D3525:=ComConveyorIO701102.o_iRequestPLCPC; 
D3526:=ComConveyorIO701102.o_iForceInportPLCPC;
D3527:=ComConveyorIO701102.o_iFolderNumberPLCPC;
D3528:=ComConveyorIO701102.o_iEmptyPLCPC;
D3530:=ComConveyorIO701102.o_iReadWriteFlagPLCPC; 
D3531:=ComConveyorIO701102.o_iDeviceStatusPLCPC; 
D3532:=ComConveyorIO701102.o_iTaskIDPLCPC; 
D3533:=ComConveyorIO701102.o_iProductIDPLCPC;
ComConveyorIO701102.i_xExportConveyor:=1;
ComConveyorIO701102.i_xExtraCondition:=ConveyorIO70159.xEmpty AND NOT ConveyorIO70159.xCWPresent AND NOT ConveyorIO701102.xCWPresent;*)
(*F5出库站台1*)
ComConveyorIO70159.i_iResponsPCPLC:=D2540; 
ComConveyorIO70159.i_iTypeInfoPCPLC:=D2541;
ComConveyorIO70159.i_iReadWriteFlagPCPLC:=D2545; 
ComConveyorIO70159.i_iTaskProcessFlagPCPLC:=D2546; 
ComConveyorIO70159.i_iCommandPCPLC:=D2547; 
ComConveyorIO70159.i_iTaskIDPCPLC:=D2548; 
DMOV(TRUE,D2549,ComConveyorIO70159.i_diDestinationDevicePCPLC); 
ComConveyorIO70159.i_iProductIDPCPLC:=D2551;
D3540:=ComConveyorIO70159.o_iRequestPLCPC; 
D3541:=ComConveyorIO70159.o_iForceInportPLCPC;
D3542:=ComConveyorIO70159.o_iFolderNumberPLCPC;
D3543:=ComConveyorIO70159.o_iEmptyPLCPC;
D3545:=ComConveyorIO70159.o_iReadWriteFlagPLCPC; 
D3546:=ComConveyorIO70159.o_iDeviceStatusPLCPC; 
D3547:=ComConveyorIO70159.o_iTaskIDPLCPC; 
D3548:=ComConveyorIO70159.o_iProductIDPLCPC;
ComConveyorIO70159.i_xExportConveyor:=1;
ComConveyorIO70159.i_xExtraCondition:=ConveyorIO701102.xEmpty AND NOT ConveyorIO70159.xCWPresent AND NOT ConveyorIO701102.xCWPresent;
(*F6出库站台1*)
ComConveyorIO701120.i_iResponsPCPLC:=D2555; 
ComConveyorIO701120.i_iTypeInfoPCPLC:=D2556;
ComConveyorIO701120.i_iReadWriteFlagPCPLC:=D2560; 
ComConveyorIO701120.i_iTaskProcessFlagPCPLC:=D2561; 
ComConveyorIO701120.i_iCommandPCPLC:=D2562; 
ComConveyorIO701120.i_iTaskIDPCPLC:=D2563; 
DMOV(TRUE,D2564,ComConveyorIO701120.i_diDestinationDevicePCPLC); 
ComConveyorIO701120.i_iProductIDPCPLC:=D2566;
D3555:=ComConveyorIO701120.o_iRequestPLCPC; 
D3556:=ComConveyorIO701120.o_iForceInportPLCPC;
D3557:=ComConveyorIO701120.o_iFolderNumberPLCPC;
D3558:=ComConveyorIO701120.o_iEmptyPLCPC;
D3560:=ComConveyorIO701120.o_iReadWriteFlagPLCPC; 
D3561:=ComConveyorIO701120.o_iDeviceStatusPLCPC; 
D3562:=ComConveyorIO701120.o_iTaskIDPLCPC; 
D3563:=ComConveyorIO701120.o_iProductIDPLCPC;
ComConveyorIO701120.i_xExportConveyor:=1;
ComConveyorIO701120.i_xExtraCondition:=ConveyorIO701119.xEmpty AND NOT ConveyorIO701119.xCWPresent AND NOT ConveyorIO701120.xCWPresent;
(*
ComConveyorIO701119.i_iResponsPCPLC:=D2570; 
ComConveyorIO701119.i_iTypeInfoPCPLC:=D2571;
ComConveyorIO701119.i_iReadWriteFlagPCPLC:=D2575; 
ComConveyorIO701119.i_iTaskProcessFlagPCPLC:=D2576; 
ComConveyorIO701119.i_iCommandPCPLC:=D2577; 
ComConveyorIO701119.i_iTaskIDPCPLC:=D2578; 
DMOV(TRUE,D2579,ComConveyorIO701119.i_diDestinationDevicePCPLC); 
ComConveyorIO701119.i_iProductIDPCPLC:=D2581;
D3570:=ComConveyorIO701119.o_iRequestPLCPC; 
D3571:=ComConveyorIO701119.o_iForceInportPLCPC;
D3572:=ComConveyorIO701119.o_iFolderNumberPLCPC;
D3573:=ComConveyorIO701119.o_iEmptyPLCPC;
D3575:=ComConveyorIO701119.o_iReadWriteFlagPLCPC; 
D3576:=ComConveyorIO701119.o_iDeviceStatusPLCPC; 
D3577:=ComConveyorIO701119.o_iTaskIDPLCPC; 
D3578:=ComConveyorIO701119.o_iProductIDPLCPC;
ComConveyorIO701119.i_xExportConveyor:=1;*)
(*F1空框入库站台2*)
ComConveyorIO701105.i_iTypeInfoPCPLC:=D2616;
ComConveyorIO701105.i_iReadWriteFlagPCPLC:=D2620; 
ComConveyorIO701105.i_iTaskProcessFlagPCPLC:=D2621; 
ComConveyorIO701105.i_iCommandPCPLC:=D2622; 
ComConveyorIO701105.i_iTaskIDPCPLC:=D2623; 
DMOV(TRUE,D2624,ComConveyorIO701105.i_diDestinationDevicePCPLC); 
ComConveyorIO701105.i_iProductIDPCPLC:=D2626;
D3615:=ComConveyorIO701105.o_iRequestPLCPC; 
D3616:=ComConveyorIO701105.o_iForceInportPLCPC;
D3617:=ComConveyorIO701105.o_iFolderNumberPLCPC;
D3618:=ComConveyorIO701105.o_iEmptyPLCPC;
D3620:=ComConveyorIO701105.o_iReadWriteFlagPLCPC; 
D3621:=ComConveyorIO701105.o_iDeviceStatusPLCPC; 
D3622:=ComConveyorIO701105.o_iTaskIDPLCPC; 
D3623:=ComConveyorIO701105.o_iProductIDPLCPC;
(*F2空框入库站台1*)
ComConveyorIO70113.i_iResponsPCPLC:=D2630; 
ComConveyorIO70113.i_iTypeInfoPCPLC:=D2631;
ComConveyorIO70113.i_iReadWriteFlagPCPLC:=D2635; 
ComConveyorIO70113.i_iTaskProcessFlagPCPLC:=D2636; 
ComConveyorIO70113.i_iCommandPCPLC:=D2637; 
ComConveyorIO70113.i_iTaskIDPCPLC:=D2638; 
DMOV(TRUE,D2639,ComConveyorIO70113.i_diDestinationDevicePCPLC); 
ComConveyorIO70113.i_iProductIDPCPLC:=D2641;
D3630:=ComConveyorIO70113.o_iRequestPLCPC; 
D3631:=ComConveyorIO70113.o_iForceInportPLCPC;
D3632:=ComConveyorIO70113.o_iFolderNumberPLCPC;
D3633:=ComConveyorIO70113.o_iEmptyPLCPC;
D3635:=ComConveyorIO70113.o_iReadWriteFlagPLCPC; 
D3636:=ComConveyorIO70113.o_iDeviceStatusPLCPC; 
D3637:=ComConveyorIO70113.o_iTaskIDPLCPC; 
D3638:=ComConveyorIO70113.o_iProductIDPLCPC;
(*F2空框入库站台2*)
ComConveyorIO701106.i_iResponsPCPLC:=D2645; 
ComConveyorIO701106.i_iTypeInfoPCPLC:=D2646;
ComConveyorIO701106.i_iReadWriteFlagPCPLC:=D2650; 
ComConveyorIO701106.i_iTaskProcessFlagPCPLC:=D2651; 
ComConveyorIO701106.i_iCommandPCPLC:=D2652; 
ComConveyorIO701106.i_iTaskIDPCPLC:=D2653; 
DMOV(TRUE,D2654,ComConveyorIO701106.i_diDestinationDevicePCPLC); 
ComConveyorIO701106.i_iProductIDPCPLC:=D2656;
D3645:=ComConveyorIO701106.o_iRequestPLCPC; 
D3646:=ComConveyorIO701106.o_iForceInportPLCPC;
D3647:=ComConveyorIO701106.o_iFolderNumberPLCPC;
D3648:=ComConveyorIO701106.o_iEmptyPLCPC;
D3650:=ComConveyorIO701106.o_iReadWriteFlagPLCPC; 
D3651:=ComConveyorIO701106.o_iDeviceStatusPLCPC; 
D3652:=ComConveyorIO701106.o_iTaskIDPLCPC; 
D3653:=ComConveyorIO701106.o_iProductIDPLCPC;
(*F1,2入库前主路分流站台*)
ComConveyorIO70114.i_iResponsPCPLC:=D2660; 
ComConveyorIO70114.i_iTypeInfoPCPLC:=D2661;
ComConveyorIO70114.i_iReadWriteFlagPCPLC:=D2665; 
ComConveyorIO70114.i_iTaskProcessFlagPCPLC:=D2666; 
ComConveyorIO70114.i_iCommandPCPLC:=D2667; 
ComConveyorIO70114.i_iTaskIDPCPLC:=D2668; 
DMOV(TRUE,D2669,ComConveyorIO70114.i_diDestinationDevicePCPLC); 
ComConveyorIO70114.i_iProductIDPCPLC:=D2671;
D3660:=ComConveyorIO70114.o_iRequestPLCPC; 
D3661:=ComConveyorIO70114.o_iForceInportPLCPC;
D3662:=ComConveyorIO70114.o_iFolderNumberPLCPC;
D3663:=ComConveyorIO70114.o_iEmptyPLCPC;
D3665:=ComConveyorIO70114.o_iReadWriteFlagPLCPC; 
D3666:=ComConveyorIO70114.o_iDeviceStatusPLCPC; 
D3667:=ComConveyorIO70114.o_iTaskIDPLCPC; 
D3668:=ComConveyorIO70114.o_iProductIDPLCPC;
ComConveyorIO70116.i_iTypeInfoPCPLC:=D2691;
ComConveyorIO70116.i_iReadWriteFlagPCPLC:=D2695; 
ComConveyorIO70116.i_iTaskProcessFlagPCPLC:=D2696; 
ComConveyorIO70116.i_iCommandPCPLC:=D2697; 
ComConveyorIO70116.i_iTaskIDPCPLC:=D2698; 
DMOV(TRUE,D2699,ComConveyorIO70116.i_diDestinationDevicePCPLC); 
ComConveyorIO70116.i_iProductIDPCPLC:=D2701;
D3690:=ComConveyorIO70116.o_iRequestPLCPC; 
D3691:=ComConveyorIO70116.o_iForceInportPLCPC;
D3692:=ComConveyorIO70116.o_iFolderNumberPLCPC;
D3693:=ComConveyorIO70116.o_iEmptyPLCPC;
D3695:=ComConveyorIO70116.o_iReadWriteFlagPLCPC; 
D3696:=ComConveyorIO70116.o_iDeviceStatusPLCPC; 
D3697:=ComConveyorIO70116.o_iTaskIDPLCPC; 
D3698:=ComConveyorIO70116.o_iProductIDPLCPC;
ComConveyorIO70119.i_iResponsPCPLC:=D2705; 
ComConveyorIO70119.i_iTypeInfoPCPLC:=D2706;
ComConveyorIO70119.i_iReadWriteFlagPCPLC:=D2710; 
ComConveyorIO70119.i_iTaskProcessFlagPCPLC:=D2711; 
ComConveyorIO70119.i_iCommandPCPLC:=D2712; 
ComConveyorIO70119.i_iTaskIDPCPLC:=D2713; 
DMOV(TRUE,D2714,ComConveyorIO70119.i_diDestinationDevicePCPLC); 
ComConveyorIO70119.i_iProductIDPCPLC:=D2716;
D3705:=ComConveyorIO70119.o_iRequestPLCPC; 
D3706:=ComConveyorIO70119.o_iForceInportPLCPC;
D3707:=ComConveyorIO70119.o_iFolderNumberPLCPC;
D3708:=ComConveyorIO70119.o_iEmptyPLCPC;
D3710:=ComConveyorIO70119.o_iReadWriteFlagPLCPC; 
D3711:=ComConveyorIO70119.o_iDeviceStatusPLCPC; 
D3712:=ComConveyorIO70119.o_iTaskIDPLCPC; 
D3713:=ComConveyorIO70119.o_iProductIDPLCPC;
ComConveyorIO70120.i_iResponsPCPLC:=D2720; 
ComConveyorIO70120.i_iTypeInfoPCPLC:=D2721;
ComConveyorIO70120.i_iReadWriteFlagPCPLC:=D2725; 
ComConveyorIO70120.i_iTaskProcessFlagPCPLC:=D2726; 
ComConveyorIO70120.i_iCommandPCPLC:=D2727; 
ComConveyorIO70120.i_iTaskIDPCPLC:=D2728; 
DMOV(TRUE,D2729,ComConveyorIO70120.i_diDestinationDevicePCPLC); 
ComConveyorIO70120.i_iProductIDPCPLC:=D2731;
D3720:=ComConveyorIO70120.o_iRequestPLCPC; 
D3721:=ComConveyorIO70120.o_iForceInportPLCPC;
D3722:=ComConveyorIO70120.o_iFolderNumberPLCPC;
D3723:=ComConveyorIO70120.o_iEmptyPLCPC;
D3725:=ComConveyorIO70120.o_iReadWriteFlagPLCPC; 
D3726:=ComConveyorIO70120.o_iDeviceStatusPLCPC; 
D3727:=ComConveyorIO70120.o_iTaskIDPLCPC; 
D3728:=ComConveyorIO70120.o_iProductIDPLCPC;
ComConveyorIO701107.i_iResponsPCPLC:=D2735; 
ComConveyorIO701107.i_iTypeInfoPCPLC:=D2736;
ComConveyorIO701107.i_iReadWriteFlagPCPLC:=D2740; 
ComConveyorIO701107.i_iTaskProcessFlagPCPLC:=D2741; 
ComConveyorIO701107.i_iCommandPCPLC:=D2742; 
ComConveyorIO701107.i_iTaskIDPCPLC:=D2743; 
DMOV(TRUE,D2744,ComConveyorIO701107.i_diDestinationDevicePCPLC); 
ComConveyorIO701107.i_iProductIDPCPLC:=D2746;
D3735:=ComConveyorIO701107.o_iRequestPLCPC; 
D3736:=ComConveyorIO701107.o_iForceInportPLCPC;
D3737:=ComConveyorIO701107.o_iFolderNumberPLCPC;
D3738:=ComConveyorIO701107.o_iEmptyPLCPC;
D3740:=ComConveyorIO701107.o_iReadWriteFlagPLCPC; 
D3741:=ComConveyorIO701107.o_iDeviceStatusPLCPC; 
D3742:=ComConveyorIO701107.o_iTaskIDPLCPC; 
D3743:=ComConveyorIO701107.o_iProductIDPLCPC;
ComConveyorIO70121.i_iResponsPCPLC:=D2750; 
ComConveyorIO70121.i_iTypeInfoPCPLC:=D2751;
ComConveyorIO70121.i_iReadWriteFlagPCPLC:=D2755; 
ComConveyorIO70121.i_iTaskProcessFlagPCPLC:=D2756; 
ComConveyorIO70121.i_iCommandPCPLC:=D2757; 
ComConveyorIO70121.i_iTaskIDPCPLC:=D2758; 
DMOV(TRUE,D2759,ComConveyorIO70121.i_diDestinationDevicePCPLC); 
ComConveyorIO70121.i_iProductIDPCPLC:=D2761;
D3750:=ComConveyorIO70121.o_iRequestPLCPC; 
D3751:=ComConveyorIO70121.o_iForceInportPLCPC;
D3752:=ComConveyorIO70121.o_iFolderNumberPLCPC;
D3753:=ComConveyorIO70121.o_iEmptyPLCPC;
D3755:=ComConveyorIO70121.o_iReadWriteFlagPLCPC; 
D3756:=ComConveyorIO70121.o_iDeviceStatusPLCPC; 
D3757:=ComConveyorIO70121.o_iTaskIDPLCPC; 
D3758:=ComConveyorIO70121.o_iProductIDPLCPC;
ComConveyorIO701108.i_iResponsPCPLC:=D2765; 
ComConveyorIO701108.i_iTypeInfoPCPLC:=D2766;
ComConveyorIO701108.i_iReadWriteFlagPCPLC:=D2770; 
ComConveyorIO701108.i_iTaskProcessFlagPCPLC:=D2771; 
ComConveyorIO701108.i_iCommandPCPLC:=D2772; 
ComConveyorIO701108.i_iTaskIDPCPLC:=D2773; 
DMOV(TRUE,D2774,ComConveyorIO701108.i_diDestinationDevicePCPLC); 
ComConveyorIO701108.i_iProductIDPCPLC:=D2776;
D3765:=ComConveyorIO701108.o_iRequestPLCPC; 
D3766:=ComConveyorIO701108.o_iForceInportPLCPC;
D3767:=ComConveyorIO701108.o_iFolderNumberPLCPC;
D3768:=ComConveyorIO701108.o_iEmptyPLCPC;
D3770:=ComConveyorIO701108.o_iReadWriteFlagPLCPC; 
D3771:=ComConveyorIO701108.o_iDeviceStatusPLCPC; 
D3772:=ComConveyorIO701108.o_iTaskIDPLCPC; 
D3773:=ComConveyorIO701108.o_iProductIDPLCPC;
ComConveyorIO70122.i_iResponsPCPLC:=D2780; 
ComConveyorIO70122.i_iTypeInfoPCPLC:=D2781;
ComConveyorIO70122.i_iReadWriteFlagPCPLC:=D2785; 
ComConveyorIO70122.i_iTaskProcessFlagPCPLC:=D2786; 
ComConveyorIO70122.i_iCommandPCPLC:=D2787; 
ComConveyorIO70122.i_iTaskIDPCPLC:=D2788; 
DMOV(TRUE,D2789,ComConveyorIO70122.i_diDestinationDevicePCPLC); 
ComConveyorIO70122.i_iProductIDPCPLC:=D2791;
D3780:=ComConveyorIO70122.o_iRequestPLCPC; 
D3781:=ComConveyorIO70122.o_iForceInportPLCPC;
D3782:=ComConveyorIO70122.o_iFolderNumberPLCPC;
D3783:=ComConveyorIO70122.o_iEmptyPLCPC;
D3785:=ComConveyorIO70122.o_iReadWriteFlagPLCPC; 
D3786:=ComConveyorIO70122.o_iDeviceStatusPLCPC; 
D3787:=ComConveyorIO70122.o_iTaskIDPLCPC; 
D3788:=ComConveyorIO70122.o_iProductIDPLCPC;
ComConveyorIO70124.i_iResponsPCPLC:=D2795; 
ComConveyorIO70124.i_iTypeInfoPCPLC:=D2796;
ComConveyorIO70124.i_iReadWriteFlagPCPLC:=D2800; 
ComConveyorIO70124.i_iTaskProcessFlagPCPLC:=D2801; 
ComConveyorIO70124.i_iCommandPCPLC:=D2802; 
ComConveyorIO70124.i_iTaskIDPCPLC:=D2803; 
DMOV(TRUE,D2804,ComConveyorIO70124.i_diDestinationDevicePCPLC); 
ComConveyorIO70124.i_iProductIDPCPLC:=D2806;
D3795:=ComConveyorIO70124.o_iRequestPLCPC; 
D3796:=ComConveyorIO70124.o_iForceInportPLCPC;
D3797:=ComConveyorIO70124.o_iFolderNumberPLCPC;
D3798:=ComConveyorIO70124.o_iEmptyPLCPC;
D3800:=ComConveyorIO70124.o_iReadWriteFlagPLCPC; 
D3801:=ComConveyorIO70124.o_iDeviceStatusPLCPC; 
D3802:=ComConveyorIO70124.o_iTaskIDPLCPC; 
D3803:=ComConveyorIO70124.o_iProductIDPLCPC;
ComConveyorIO70127.i_iResponsPCPLC:=D2810; 
ComConveyorIO70127.i_iTypeInfoPCPLC:=D2811;
ComConveyorIO70127.i_iReadWriteFlagPCPLC:=D2815; 
ComConveyorIO70127.i_iTaskProcessFlagPCPLC:=D2816; 
ComConveyorIO70127.i_iCommandPCPLC:=D2817; 
ComConveyorIO70127.i_iTaskIDPCPLC:=D2818; 
DMOV(TRUE,D2819,ComConveyorIO70127.i_diDestinationDevicePCPLC); 
ComConveyorIO70127.i_iProductIDPCPLC:=D2821;
D3810:=ComConveyorIO70127.o_iRequestPLCPC; 
D3811:=ComConveyorIO70127.o_iForceInportPLCPC;
D3812:=ComConveyorIO70127.o_iFolderNumberPLCPC;
D3813:=ComConveyorIO70127.o_iEmptyPLCPC;
D3815:=ComConveyorIO70127.o_iReadWriteFlagPLCPC; 
D3816:=ComConveyorIO70127.o_iDeviceStatusPLCPC; 
D3817:=ComConveyorIO70127.o_iTaskIDPLCPC; 
D3818:=ComConveyorIO70127.o_iProductIDPLCPC;
ComConveyorIO70128.i_iResponsPCPLC:=D2825; 
ComConveyorIO70128.i_iTypeInfoPCPLC:=D2826;
ComConveyorIO70128.i_iReadWriteFlagPCPLC:=D2830; 
ComConveyorIO70128.i_iTaskProcessFlagPCPLC:=D2831; 
ComConveyorIO70128.i_iCommandPCPLC:=D2832; 
ComConveyorIO70128.i_iTaskIDPCPLC:=D2833; 
DMOV(TRUE,D2834,ComConveyorIO70128.i_diDestinationDevicePCPLC); 
ComConveyorIO70128.i_iProductIDPCPLC:=D2836;
D3825:=ComConveyorIO70128.o_iRequestPLCPC; 
D3826:=ComConveyorIO70128.o_iForceInportPLCPC;
D3827:=ComConveyorIO70128.o_iFolderNumberPLCPC;
D3828:=ComConveyorIO70128.o_iEmptyPLCPC;
D3830:=ComConveyorIO70128.o_iReadWriteFlagPLCPC; 
D3831:=ComConveyorIO70128.o_iDeviceStatusPLCPC; 
D3832:=ComConveyorIO70128.o_iTaskIDPLCPC; 
D3833:=ComConveyorIO70128.o_iProductIDPLCPC;
ComConveyorIO701109.i_iResponsPCPLC:=D2840; 
ComConveyorIO701109.i_iTypeInfoPCPLC:=D2841;
ComConveyorIO701109.i_iReadWriteFlagPCPLC:=D2845; 
ComConveyorIO701109.i_iTaskProcessFlagPCPLC:=D2846; 
ComConveyorIO701109.i_iCommandPCPLC:=D2847; 
ComConveyorIO701109.i_iTaskIDPCPLC:=D2848; 
DMOV(TRUE,D2849,ComConveyorIO701109.i_diDestinationDevicePCPLC); 
ComConveyorIO701109.i_iProductIDPCPLC:=D2851;
D3840:=ComConveyorIO701109.o_iRequestPLCPC; 
D3841:=ComConveyorIO701109.o_iForceInportPLCPC;
D3842:=ComConveyorIO701109.o_iFolderNumberPLCPC;
D3843:=ComConveyorIO701109.o_iEmptyPLCPC;
D3845:=ComConveyorIO701109.o_iReadWriteFlagPLCPC; 
D3846:=ComConveyorIO701109.o_iDeviceStatusPLCPC; 
D3847:=ComConveyorIO701109.o_iTaskIDPLCPC; 
D3848:=ComConveyorIO701109.o_iProductIDPLCPC;
ComConveyorIO70129.i_iResponsPCPLC:=D2855; 
ComConveyorIO70129.i_iTypeInfoPCPLC:=D2856;
ComConveyorIO70129.i_iReadWriteFlagPCPLC:=D2860; 
ComConveyorIO70129.i_iTaskProcessFlagPCPLC:=D2861; 
ComConveyorIO70129.i_iCommandPCPLC:=D2862; 
ComConveyorIO70129.i_iTaskIDPCPLC:=D2863; 
DMOV(TRUE,D2864,ComConveyorIO70129.i_diDestinationDevicePCPLC); 
ComConveyorIO70129.i_iProductIDPCPLC:=D2866;
D3855:=ComConveyorIO70129.o_iRequestPLCPC; 
D3856:=ComConveyorIO70129.o_iForceInportPLCPC;
D3857:=ComConveyorIO70129.o_iFolderNumberPLCPC;
D3858:=ComConveyorIO70129.o_iEmptyPLCPC;
D3860:=ComConveyorIO70129.o_iReadWriteFlagPLCPC; 
D3861:=ComConveyorIO70129.o_iDeviceStatusPLCPC; 
D3862:=ComConveyorIO70129.o_iTaskIDPLCPC;
D3863:=ComConveyorIO70129.o_iProductIDPLCPC;
ComConveyorIO701110.i_iResponsPCPLC:=D2870; 
ComConveyorIO701110.i_iTypeInfoPCPLC:=D2871;
ComConveyorIO701110.i_iReadWriteFlagPCPLC:=D2875; 
ComConveyorIO701110.i_iTaskProcessFlagPCPLC:=D2876; 
ComConveyorIO701110.i_iCommandPCPLC:=D2877; 
ComConveyorIO701110.i_iTaskIDPCPLC:=D2878; 
DMOV(TRUE,D2879,ComConveyorIO701110.i_diDestinationDevicePCPLC); 
ComConveyorIO701110.i_iProductIDPCPLC:=D2881;
D3870:=ComConveyorIO701110.o_iRequestPLCPC; 
D3871:=ComConveyorIO701110.o_iForceInportPLCPC;
D3872:=ComConveyorIO701110.o_iFolderNumberPLCPC;
D3873:=ComConveyorIO701110.o_iEmptyPLCPC;
D3875:=ComConveyorIO701110.o_iReadWriteFlagPLCPC; 
D3876:=ComConveyorIO701110.o_iDeviceStatusPLCPC; 
D3877:=ComConveyorIO701110.o_iTaskIDPLCPC; 
D3878:=ComConveyorIO701110.o_iProductIDPLCPC;

(*OCV2分拣通信程序*)
SortCommunication70210(ConveyorIO:=ConveyorIO70173,SortCommunicationIO:= SortCommunicationIO70210 ,FanucRobotIO:= RobotIO70210,ServoIO:=ServoIO1);
SortCommunicationIO70210 .i_iResponsPCPLC:=D2705;
SortCommunicationIO70210 .i_iInfoWriteDone:=D2706;
SortCommunicationIO70210 .i_iSortDoneAknPCPLC:=D2707;
D3705:=SortCommunicationIO70210 .o_iRequestPLCPC;(*有料请求*)
D3706:=SortCommunicationIO70210 .o_iSortDonePLCPC;(*分拣完成信号*)
FOR Z0:=0 TO 127 BY 1 DO
	SortCommunicationIO70210 .i_arriBatteryStatus[Z0+1]:=D2708Z0;
END_FOR;
SortCommunicationIO70210 .i_xSortOver:=X66;
RobotIO70210.i_xPickOver:=X118;(*机器人给的取货完成*)
RobotIO70210.i_xPutOver:=X11A;(*机器人给的放货完成*)
Y3B4:=RobotIO70210.o_xSortStart;(*给机器人的开始启动*)
Y3A3:=RobotIO70210.o_xColumn[0];(*给机器人的行号*)
Y3B5:=RobotIO70210.o_xColumn[1];
Y3A4:=RobotIO70210.o_xColumn[2];
Y3B7:=RobotIO70210.o_xColumn[3];
Y3A6:=RobotIO70210.o_xRow[0];(*给机器人的列号*)
Y3A8:=RobotIO70210.o_xRow[1];
Y3A7:=RobotIO70210.o_xRow[2];
Y3A5:=RobotIO70210.o_xRow[3];
Y3B6:=RobotIO70210.o_xPutNumber[0];(*给机器人的放料位置*)
Y3A2:=RobotIO70210.o_xPutNumber[1];
Y3A1:=RobotIO70210.o_xPutNumber[2];
Y3B8:=RobotIO70210.o_xPutNumber[3];
Y2A1:=RobotIO70210.o_xCatchCylinder;
RobotIO70210.i_xBatteryDetect[3]:=X7F;
RobotIO70210.i_xBatteryDetect[2]:=XF4;
RobotIO70210.i_xBatteryDetect[1]:=XF6;
RobotIO70210.i_xBatteryDetect[0]:=XF9;
RobotIO70210.i_xProtect[0]:=X7E;
RobotIO70210.i_xProtect[1]:=XE5;
RobotIO70210.i_xProtect[2]:=XE4;
RobotIO70210.i_xProtect[3]:=XFB;

(*OCV2分拣排废线调用*)
Servo1(ServoIO:=ServoIO1 ,xAuto:=g_xAuto ,xManual:= g_xManual );
Y380:=ServoIO1.xPLCReady;
ServoIO1.xQD75Error1:=X388;					ServoIO1.xQD75Error2:=X389;		ServoIO1.xQD75Error3:=X38A;		ServoIO1.xQD75Error4:=X38B;
ServoIO1.xQD75Busy1:=X38C;				ServoIO1.xQD75Busy2:=X38D;		ServoIO1.xQD75Busy3:=X38E;		ServoIO1.xQD75Busy4:=X38F;
ServoIO1.xQD75LocateDone1:=X394;	ServoIO1.xQD75LocateDone2:=X395;	ServoIO1.xQD75LocateDone3:=X396;	ServoIO1.xQD75LocateDone4:=X397;
Y390:=ServoIO1.xQD75LocateStart1;	Y391:=ServoIO1.xQD75LocateStart2;	Y392:=ServoIO1.xQD75LocateStart3;	Y393:=ServoIO1.xQD75LocateStart4;
(*OCV2刹车控制，懒得单独写，就这样了*)
Y2CB:=ServoIO1.xQD75LocateStart1;	Y2CF:=ServoIO1.xQD75LocateStart2;	Y2D1:=ServoIO1.xQD75LocateStart3;	Y2D3:=ServoIO1.xQD75LocateStart4;
DMOV(TRUE,U38\G800,ServoIO1.diQD75CurrentPos1);(*当前位置*)	DMOV(TRUE,U38\G900,ServoIO1.diQD75CurrentPos2);(*当前位置*)
DMOV(TRUE,U38\G1000,ServoIO1.diQD75CurrentPos3);(*当前位置*)	DMOV(TRUE,U38\G1100,ServoIO1.diQD75CurrentPos4);(*当前位置*)
U38\G1502:=ServoIO1.iReset1;(*轴出错复位*)	U38\G1602:=ServoIO1.iReset2;(*轴出错复位*)
U38\G1702:=ServoIO1.iReset3;(*轴出错复位*)	U38\G1802:=ServoIO1.iReset4;(*轴出错复位*)
U38\G1500:=ServoIO1.iLocateStartNumber1;(*目标地址*)	U38\G1600:=ServoIO1.iLocateStartNumber2;(*目标地址*)
U38\G1700:=ServoIO1.iLocateStartNumber3;(*目标地址*)	U38\G1800:=ServoIO1.iLocateStartNumber4;(*目标地址*)

(*OCV3分拣通信程序*)
SortCommunication70184(ConveyorIO:=ConveyorIO70184,SortCommunicationIO:= SortCommunicationIO70184 ,FanucRobotIO:= RobotIO70184,ServoIO:=ServoIO2);
SortCommunicationIO70184 .i_iResponsPCPLC:=D2845;
SortCommunicationIO70184 .i_iInfoWriteDone:=D2846;
SortCommunicationIO70184 .i_iSortDoneAknPCPLC:=D2847;
D3845:=SortCommunicationIO70184 .o_iRequestPLCPC;(*有料请求*)
D3846:=SortCommunicationIO70184 .o_iSortDonePLCPC;(*分拣完成信号*)
FOR Z1:=0 TO 127 BY 1 DO
	SortCommunicationIO70184 .i_arriBatteryStatus[Z1+1]:=D2848Z1;
END_FOR;
(*_SortCommunicationIO70184 .i_xSortOver:=X66;这个是放行按钮，没有按钮之前先屏蔽_*)
RobotIO70184.i_xPickOver:=X129;(*机器人给的取货完成*)
RobotIO70184.i_xPutOver:=X12A;(*机器人给的放货完成*)
Y3B9:=RobotIO70184.o_xSortStart;(*给机器人的开始启动*)
Y3AF:=RobotIO70184.o_xColumn[0];(*给机器人的行号*)
Y3AA:=RobotIO70184.o_xColumn[1];
Y3B0:=RobotIO70184.o_xColumn[2];
Y3B2:=RobotIO70184.o_xColumn[3];
Y3AD:=RobotIO70184.o_xRow[0];(*给机器人的列号*)
Y3BA:=RobotIO70184.o_xRow[1];
Y3AB:=RobotIO70184.o_xRow[2];
Y3B1:=RobotIO70184.o_xRow[3];
Y3BB:=RobotIO70184.o_xPutNumber[0];(*给机器人的放料位置*)
Y3AE:=RobotIO70184.o_xPutNumber[1];
Y3AC:=RobotIO70184.o_xPutNumber[2];
Y3B3:=RobotIO70184.o_xPutNumber[3];
Y2D7:=RobotIO70184.o_xCatchCylinder;
RobotIO70184.i_xBatteryDetect[3]:=X10C;
RobotIO70184.i_xBatteryDetect[2]:=X10B;
RobotIO70184.i_xBatteryDetect[1]:=X10A;
RobotIO70184.i_xBatteryDetect[0]:=X109;
RobotIO70184.i_xProtect[0]:=X100;
RobotIO70184.i_xProtect[1]:=X101;
RobotIO70184.i_xProtect[2]:=X102;
RobotIO70184.i_xProtect[3]:=X103;

(*OCV3分拣排废线调用*)
Servo2(ServoIO:=ServoIO2 ,xAuto:=g_xAuto ,xManual:= g_xManual );
Y3E0:=ServoIO2.xPLCReady;
ServoIO2.xQD75Error1:=X3E8;					ServoIO2.xQD75Error2:=X3E9;		ServoIO2.xQD75Error3:=X3EA;		ServoIO2.xQD75Error4:=X3EB;
ServoIO2.xQD75Busy1:=X3EC;				ServoIO2.xQD75Busy2:=X3ED;		ServoIO2.xQD75Busy3:=X3EE;		ServoIO2.xQD75Busy4:=X3EF;
ServoIO2.xQD75LocateDone1:=X3F4;	ServoIO2.xQD75LocateDone2:=X3F5;	ServoIO2.xQD75LocateDone3:=X3F6;	ServoIO2.xQD75LocateDone4:=X3F7;
Y3F0:=ServoIO2.xQD75LocateStart1;	Y3F1:=ServoIO2.xQD75LocateStart2;	Y3F2:=ServoIO2.xQD75LocateStart3;	Y3F3:=ServoIO2.xQD75LocateStart4;
(*OCV3刹车控制，懒得单独写，就这样了*)
Y2D5:=ServoIO2.xQD75LocateStart1;	Y2D9:=ServoIO2.xQD75LocateStart2;	Y2DB:=ServoIO2.xQD75LocateStart3;	Y2DD:=ServoIO2.xQD75LocateStart4;
(*
DMOV(TRUE,U3E\G800,ServoIO2.diQD75CurrentPos1);(*当前位置*)(*	DMOV(TRUE,U3E\G900,ServoIO2.diQD75CurrentPos2);(*当前位置*)(*
DMOV(TRUE,U3E\G1000,ServoIO2.diQD75CurrentPos3);(*当前位置*)	(*DMOV(TRUE,U3E\G1100,ServoIO2.diQD75CurrentPos4);(*当前位置*)(*
U3E\G1502:=ServoIO2.iReset1;(*轴出错复位*)(*	U3E\G1602:=ServoIO2.iReset2;(*轴出错复位*)(*
U3E\G1702:=ServoIO2.iReset3;(*轴出错复位*)(*	U3E\G1802:=ServoIO2.iReset4;(*轴出错复位*)(*
U3E\G1500:=ServoIO2.iLocateStartNumber1;(*目标地址*)(*	U3E\G1600:=ServoIO2.iLocateStartNumber2;(*目标地址*)(*
U3E\G1700:=ServoIO2.iLocateStartNumber3;(*目标地址*)(*	U3E\G1800:=ServoIO2.iLocateStartNumber4;(*目标地址*)


(*线体信息传递*)
(*1#入库*)
ConveyorIO70195.diDesConveyorIn:= ConveyorIO70190.diDesConveyorOut;
ConveyorIO70196.diDesConveyorIn:= ConveyorIO70190.diDesConveyorOut;
ConveyorIO70146.diDesConveyorIn:= ConveyorIO70195.diDesConveyorOut;
ConveyorIO70147.diDesConveyorIn:= ConveyorIO70196.diDesConveyorOut;
ConveyorIO70195.iTaskIDIn:= ConveyorIO70190.iTaskIDOut;
ConveyorIO70196.iTaskIDIn:= ConveyorIO70190.iTaskIDOut;
ConveyorIO70146.iTaskIDIn:= ConveyorIO70195.iTaskIDOut;
ConveyorIO70147.iTaskIDIn:= ConveyorIO70196.iTaskIDOut;
ConveyorIO70195.iProductCategoryIn:= ConveyorIO70190.iProductCategoryOut;
ConveyorIO70196.iProductCategoryIn:= ConveyorIO70190.iProductCategoryOut;
ConveyorIO70146.iProductCategoryIn:= ConveyorIO70195.iProductCategoryOut;
ConveyorIO70147.iProductCategoryIn:= ConveyorIO70196.iProductCategoryOut;
(*2#入库*)
ConveyorIO70199.diDesConveyorIn:= ConveyorIO70192.diDesConveyorOut;
ConveyorIO701100.diDesConveyorIn:= ConveyorIO70192.diDesConveyorOut;
ConveyorIO70154.diDesConveyorIn:= ConveyorIO70199.diDesConveyorOut;
ConveyorIO70155.diDesConveyorIn:= ConveyorIO701100.diDesConveyorOut;
ConveyorIO70199.iTaskIDIn:= ConveyorIO70192.iTaskIDOut;
ConveyorIO701100.iTaskIDIn:= ConveyorIO70192.iTaskIDOut;
ConveyorIO70154.iTaskIDIn:= ConveyorIO70199.iTaskIDOut;
ConveyorIO70155.iTaskIDIn:= ConveyorIO701100.iTaskIDOut;
ConveyorIO70199.iProductCategoryIn:= ConveyorIO70192.iProductCategoryOut;
ConveyorIO701100.iProductCategoryIn:= ConveyorIO70192.iProductCategoryOut;
ConveyorIO70154.iProductCategoryIn:= ConveyorIO70199.iProductCategoryOut;
ConveyorIO70155.iProductCategoryIn:= ConveyorIO701100.iProductCategoryOut;
(*3#入库*)
ConveyorIO701103.diDesConveyorIn:= ConveyorIO70194.diDesConveyorOut;
ConveyorIO701104.diDesConveyorIn:= ConveyorIO70194.diDesConveyorOut;
ConveyorIO70162.diDesConveyorIn:= ConveyorIO701103.diDesConveyorOut;
ConveyorIO70163.diDesConveyorIn:= ConveyorIO701104.diDesConveyorOut;
ConveyorIO701103.iTaskIDIn:= ConveyorIO70194.iTaskIDOut;
ConveyorIO701104.iTaskIDIn:= ConveyorIO70194.iTaskIDOut;
ConveyorIO70162.iTaskIDIn:= ConveyorIO701103.iTaskIDOut;
ConveyorIO70163.iTaskIDIn:= ConveyorIO701104.iTaskIDOut;
ConveyorIO701103.iProductCategoryIn:= ConveyorIO70194.iProductCategoryOut;
ConveyorIO701104.iProductCategoryIn:= ConveyorIO70194.iProductCategoryOut;
ConveyorIO70162.iProductCategoryIn:= ConveyorIO701103.iProductCategoryOut;
ConveyorIO70163.iProductCategoryIn:= ConveyorIO701104.iProductCategoryOut;
(*自动*)
(*安全通道*)
ConveyorIO70101.xLoad:=X159;
m_x60LoadRequest:=ConveyorIO70101.xEmpty;
ConveyorIO70101.xUnload:=ConveyorIO70102.xEmpty ;
ConveyorIO70102.xLoad:=ConveyorIO70101.xNextRun;
ConveyorIO70102.xUnload:=ConveyorIO70103.xEmpty;
ConveyorIO70103.xLoad:=ConveyorIO70102.xNextRun;
ConveyorIO70103.xUnload:=ConveyorIO70104.xEmpty;
SwitchIO70301.xEntryEnable:=ConveyorIO70103.xNextRun;
SwitchIo70301.xSwithEnable:=1;
SwitchIO70301.xExitEnable:=ConveyorIO70106.xEmpty AND LifterIO70207.iCurrentPos=2 AND LifterIO70207.xPresentDetect2;
(*提升机*)
LifterIO70207.xMDIExe:=NOT (ConveyorIO70106.xError OR ConveyorIO70105.xError OR ConveyorIO70140.xError);
IF ConveyorIO70106.xEmpty THEN
	LifterIO70207.iDestinationPos:=2;
ELSE
	LifterIO70207.iDestinationPos:=1;
END_IF;
ConveyorIO70106.xLoad:=ConveyorIO70105.xNextRun;
ConveyorIO70106.xUnload:=ConveyorIO70140.xEmpty AND ConveyorIO70140_1.xEmpty AND LifterIO70207.iCurrentPos=1 AND LifterIO70207.xPresentDetect1;
ConveyorIO70140_1.xLoad:=ConveyorIO70106.xNextRun;
ConveyorIO70140_1.xUnload:=ConveyorIO70140.xEmpty (*AND ConveyorIO70140_1.diDesConveyor=70140*) AND ComConveyorIO70104.i_iResponsPCPLC=2;
FolderIO70201.i_xEntryEnable:=ConveyorIO70140_1.xNextRun;
ConveyorIO70106.xUnloadCCW:=1;

(*rgv输送*)
(*1#入库*)
SwitchIO70311.xSwithEnable:=1;
(*根据目标地址选择顶升移载下料的方向*)
IF M22 THEN
	ConveyorIO70144.diDesConveyor:=70196;
	D3045:=0;
END_IF;
IF M23 THEN(*屏蔽叠盘机*)
	m_xFolder70201Atuo:=0;
	ConveyorIO70140.xLoad:=ConveyorIO70106.xNextRun;
	FolderIO70201.o_xExitPremit:=NOT ConveyorIO70140.xEmpty;
END_IF;	
ConveyorIO70145.xUnload:=ConveyorIO70144.xEmpty;
SwitchIO70311.xEntryEnable:=ConveyorIO70145.xNextRun;
SwitchIO70311.xExitEnable:=(ConveyorIO70195.xEmpty AND (ConveyorIO70144.diDesConveyor=70195 OR ConveyorIO70144.diDesConveyor=70146))
													OR (ConveyorIO70196.xEmpty AND (ConveyorIO70144.diDesConveyor=70196 OR ConveyorIO70144.diDesConveyor=70147));
ConveyorIO70190.xUnloadCCW:=ConveyorIO70190.diDesConveyor=70196 OR ConveyorIO70190.diDesConveyor=70147;
ConveyorIO70195.xLoad:=ConveyorIO70190.xNextRun AND (ConveyorIO70144.diDesConveyor=70195 OR ConveyorIO70144.diDesConveyor=70146);
ConveyorIO70195.xUnload:=ConveyorIO70146.xEmpty  AND ConveyorIO70195.diDesConveyor=70146;
ConveyorIO70146.xLoad:=ConveyorIO70195.xNextRun;
m_xtonConveyor70195Reset(IN:=NOT ConveyorIO70195.xCWPresent,PT:=T#10s ,Q:= ConveyorIO70195.xPutInto,ET:= m_xtonConveyor70195CurTime );
m_xtonConveyor70146Reset(IN:=NOT ConveyorIO70146.xCWPresent,PT:=T#10s ,Q:= ConveyorIO70146.xPutInto,ET:= m_xtonConveyor70146CurTime );
ConveyorIO70196.xLoad:=ConveyorIO70190.xNextRun AND (ConveyorIO70144.diDesConveyor=70196 OR ConveyorIO70144.diDesConveyor=70147);
ConveyorIO70196.xUnload:=ConveyorIO70147.xEmpty AND ConveyorIO70196.diDesConveyor=70147;
ConveyorIO70147.xLoad:=ConveyorIO70196.xNextRun;
m_xtonConveyor70196Reset(IN:=NOT ConveyorIO70196.xCWPresent,PT:=T#10s ,Q:= ConveyorIO70196.xPutInto,ET:=m_xtonConveyor70196CurTime );
m_xtonConveyor70147Reset(IN:=NOT ConveyorIO70147.xCWPresent,PT:=T#10s ,Q:= ConveyorIO70147.xPutInto,ET:= m_xtonConveyor70147CurTime);
(*1#出库*)
(*自动刷新物料状态，有料检测后10秒开始输送*)
m_xtonConveyor701115Reset(IN:=ConveyorIO701115.xCWPresent,PT:=T#10s ,Q:= ConveyorIO701115.xPutInto,ET:= m_xtonConveyor701115CurTime );
m_xtonConveyor701114Reset(IN:=ConveyorIO701114.xCWPresent,PT:=T#10s ,Q:= ConveyorIO701114.xPutInto,ET:= m_xtonConveyor701114CurTime );
ConveyorIO701114.tLoadDelay:=t#3s;
ConveyorIO701115.xUnload:=ConveyorIO701114.xEmpty;
ConveyorIO701114.xLoad:=ConveyorIO701115.xNextRun;
ConveyorIO701114.xUnload:=ConveyorIO701113.xEmpty;
SwitchIO70326.xEntryEnable:=ConveyorIO701114.xNextRun;
SwitchIO70326.xSwithEnable:=1;
SwitchIO70326.xExitEnable:=ConveyorIO701111.xEmpty;
ConveyorIO701111.xLoad:=ConveyorIO701111_1.xNextRun;
(*到达RGV接料位置*)
(*SwitchIO70316.xSwithEnable:=1;
SwitchIO70316.xExitEnable:=ConveyorIO70165_2.xEmpty AND (m_xOCV2_1LoadLock OR m_xOCV2_2LoadLock);*)(*临时程序，先用1号OVCV2，以后要做任务抢占*)
(*OCV1前顶升移载，双向电机，根据m_xOCV2_1UnloadRequest信号  改变顶升移载的出线体和入线体*)
(*SwitchIO70317.xEntryEnable:=(ConveyorIO70165_1.xNextRun AND NOT m_xOCV2_1UnloadRequest) OR m_xOCV2_1UnloadRequest;
SwitchIO70317.xSwithEnable:=(m_xOCV2_1LoadRequest  AND NOT m_xOCV2_1UnloadRequest) OR m_xOCV2_1UnloadRequest;*)(*OCV设备上料请求*)
(*SwitchIo70317.xExitEnable:=(m_xOCV2_1LoadRequest AND NOT m_xOCV2_1UnloadRequest) OR (m_xOCV2_1UnloadRequest AND COnveyorIO70166.xEmpty) ;
*)

IF M24 THEN(*屏蔽拆盘机*)
	m_xDivideFolder70204Auto:=0;
	Y335:=1;
	ConveyorIO70165_2.xload:=ConveyorIO70165_1.xNextRun;
	ConveyorIO70165_2.xUnload:=(m_xOCV2_1LoadLock OR m_xOCV2_2LoadLock) AND ConveyorIO70165.xEmpty;
	ELSE
	m_xDivideFolder70204Auto:=1;
	Y335:= ((m_xOCV2_1LoadLock OR m_xOCV2_2LoadLock) AND ConveyorIO70165_2.xNextRun) OR (M632 AND g_xManual ); (*拆盘机阻挡*)
END_IF;	
	DivideFolderIO70204.o_xExitPremit:=(m_xOCV2_1LoadLock AND ConveyorIO70165.xEmpty) OR (m_xOCV2_2LoadLock AND ConveyorIO70166.xEmpty AND ConveyorIO70165.xEmpty) ;
	DivideFolderIO70204.o_xEntryPermit:=ConveyorIO70165_1.xNextRun  AND (m_xOCV2_1LoadLock OR m_xOCV2_2LoadLock);
		DivideFolderIO70204.i_FrontConveyorNextRun:=ConveyorIO70165_1.xNextRun;
	m_xtonConveyor70164Reset(IN:=NOT ConveyorIO70164.xCWPresent,PT:=T#7s ,Q:= ConveyorIO70164.xPutInto,ET:= m_xtonConveyor70164CurTime );
m_xtonConveyor70165_1Reset(IN:=NOT ConveyorIO70164.xEmpty,PT:=T#1s ,Q:= ConveyorIO70165_1.xPutInto,ET:= m_xtonConveyor70165_1CurTime );

Y2C8:=NOT ConveyorIO70165_1.xEmpty AND NOT  X27 AND NOT X60 AND  ConveyorIO70165_2.xLoad;(*OCV2入口顶升*)

(*OCV2,3信号对接*)
m_xOCV2_1LoadRequest:=X110 AND NOT  m_Ocv2_1Forbidden ;
m_xOCV2_1UnloadRequest:=X111 ;
Y2AB:=m_xOCV2_1LoadStart OR M811;
Y2AD:=m_xOCV2_1UnloadStart OR M812;

m_xOCV2_2LoadRequest:=X112 AND NOT m_Ocv2_2Forbidden;
m_xOCV2_2UnloadRequest:=X113;
Y2AF:=m_xOCV2_2LoadStart OR M813;
Y2B1:=m_xOCV2_2UnloadStart OR M814;

m_xOCV3_1LoadRequest:=X114 AND NOT m_Ocv3_1Forbidden;
m_xOCV3_1UnloadRequest:=X115;
Y2B3:=m_xOCV3_1LoadStart OR M815;
Y2B5:=m_xOCV3_1UnloadStart OR M816;


m_xOCV3_2LoadRequest:=X116 AND NOT m_Ocv3_2Forbidden;
m_xOCV3_2UnloadRequest:=X117;
Y2B7:=m_xOCV3_2LoadStart OR M817;
Y2B9:=m_xOCV3_2UnloadStart OR M818;

m_xChoose1LoadRequest:=(M910 OR ConveyorIO70173.xEmpty) AND NOT m_Choose1Forbidden;
m_xChoose1UnLoadRequest:=M911 OR (SortCommunicationIO70210.o_xSortDone (*AND  ComConveyorIO70169.i_iResponsPCPLC=2*))  ;(*需加扫码169工位应答后放行*)

m_xChoose2LoadRequest:=M912 AND NOT m_Choose2Forbidden;
m_xChoose2UnLoadRequest:=M913;

(*———————————————OCV2———————————————*)
(*OCV2下料信号互锁，上料信号不用，因为上料信号是入口前的线体有料就可以进*)
m_xOCV2_1LoadStart:=ConveyorIO70171.xNextRun AND NOT m_xOCV2_1UnLoadLock;
m_xOCV2_1UnloadStart:=ConveyorIO70171.xEmpty AND NOT m_xOCV2_1LoadLock AND (m_xChoose1LoadLock OR m_Choose1Forbidden)
												AND NOT m_xOCV2_2LoadLock AND NOT m_xOCV2_2UnLoadLock AND ConveyorIO70167.xEmpty; 
m_xOCV2_2LoadStart:=ConveyorIO70172.xNextRun AND NOT m_xOCV2_2UnLoadLock ;
m_xOCV2_2UnloadStart:=ConveyorIO70172.xEmpty AND NOT m_xOCV2_2LoadLock AND (m_xChoose1LoadLock OR m_Choose1Forbidden)
											 AND NOT m_xOCV2_1UnLoadLock AND ConveyorIO70167.xEmpty;
m_xChoose1LoadStart:=(ConveyorIO70173.xEmpty AND NOT m_xChoose1UnLoadLock) OR M920;
m_xChoose1UnLoadStart:=(ConveyorIO70173_1.xEmpty AND NOT m_xChoose1LoadLock) OR M921 ;

(*OCV2上料信号互锁*)
set(m_xOCV2_1LoadRequest  AND  NOT m_xOCV2_1UnLoadLock  AND NOT m_xOCV2_2LoadLock,m_xOCV2_1LoadLock);
rst(NOT m_xOCV2_1LoadRequest OR M970,m_xOCV2_1LoadLock);
set(m_xOCV2_2LoadRequest AND  NOT m_xOCV2_2UnLoadLock AND NOT m_xOCV2_1LoadLock AND  NOT m_xOCV2_1UnLoadLock ,m_xOCV2_2LoadLock);
rst(NOT m_xOCV2_2LoadRequest OR M971,m_xOCV2_2LoadLock);
set(m_xChoose1LoadRequest AND NOT m_xChoose1UnLoadLock AND NOT m_xOCV2_2LoadLock,m_xChoose1LoadLock);
rst(NOT m_xChoose1LoadRequest OR M972,m_xChoose1LoadLock);

(*OCV2下料信号互锁*)
set(m_xOCV2_1UnLoadRequest AND NOT m_xOCV2_1LoadLock AND NOT m_xOCV2_2LoadLock AND NOT m_xOCV2_2UnLoadLock 
		AND (m_xChoose1LoadLock OR m_Choose1Forbidden) AND ConveyorIO70166.xEmpty,m_xOCV2_1UnLoadLock);
rst(( NOT ConveyorIO70167.xEmpty AND (NOT m_xChoose1LoadLock OR  m_Choose1Forbidden))OR M973,m_xOCV2_1UnLoadLock);
set(m_xOCV2_2UnLoadRequest AND NOT m_xOCV2_2LoadLock AND (m_xChoose1LoadLock OR m_Choose1Forbidden)  
		AND NOT m_xOCV2_1UnLoadLock AND ConveyorIO70167.xEmpty,m_xOCV2_2UnLoadLock);
rst((NOT ConveyorIO70167.xEmpty AND (NOT m_xChoose1LoadLock OR  m_Choose1Forbidden))OR M974,m_xOCV2_2UnLoadLock);
set(m_xChoose1UnloadRequest AND NOT m_xChoose1LoadLock AND ConveyorIO70167.xEmpty ,m_xChoose1UnLoadLock);
rst(NOT ConveyorIO70168_1.xEmpty OR M975,m_xChoose1UnLoadLock);
(*ocv2-1顶升和阻挡*)
Y2CA:=( ConveyorIO70165.xEmpty AND m_xOCV2_1LoadLock) (*165转171顶升*)
		OR  (m_xOCV2_1UnLoadLock  AND NOT ConveyorIO70171.xEmpty AND ConveyorIO70165.xUnLoad) 
		OR (m_xOCV2_2LoadLock AND  (ConveyorIO70165.xLoad OR ConveyorIO70165.xUnLoad)) 
		OR (m_Ocv2_1Forbidden AND (ConveyorIO70165.xLoad OR  ConveyorIO70165.xUnload) AND NOT m_xOCV2_2UnLoadLock) ;
Y336:=(m_xOCV2_1UnLoadLock AND NOT ConveyorIO70171.xEmpty  AND ConveyorIO70165.xUnLoad) 
			OR (m_xOCV2_2LoadLock AND ConveyorIO70165.xUnLoad) 
			OR (m_Ocv2_1Forbidden AND (ConveyorIO70165.xLoad OR  ConveyorIO70165.xUnload)AND NOT  m_xOCV2_2UnLoadLock) ;(*165去166阻挡*)
(*ocv2-2顶升和阻挡*)
Y2CC:=(ConveyorIO70166.xload AND m_xOCV2_2LoadLock)  (*166转OCV2-2顶升*)
			OR ((ConveyorIO70166.xLoad OR ConveyorIO70166.xUnload)  AND m_xOCV2_1UnLoadLock)
			OR ( NOT ConveyorIO70172.xEmpty AND ConveyorIO70166.xUnload  AND m_xOCV2_2UnLoadLock)
			OR (m_Ocv2_2Forbidden AND (ConveyorIO70166.xLoad OR  ConveyorIO70166.xUnload));

